// TIA Portal project "Process visualization with HMI" (V15.1) (continued)
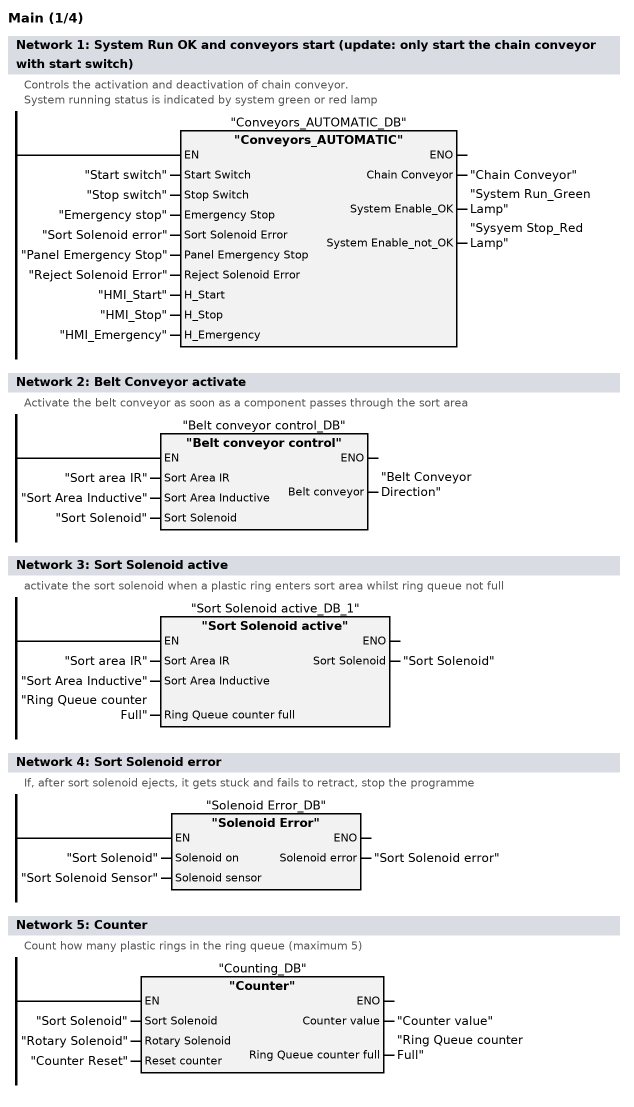
   RUNG wire#powerrail
      "Conveyors_AUTOMATIC_DB"("Start Switch" := "Start switch", "Stop Switch" := "Stop switch", "Emergency Stop" := "Emergency stop", "Sort Solenoid Error" := "Sort Solenoid error", "Panel Emergency Stop" := "Panel Emergency Stop", "Reject Solenoid Error" := "Reject Solenoid Error", H_Start := "HMI_Start", H_Stop := "HMI_Stop", H_Emergency := "HMI_Emergency", "Chain Conveyor" => "Chain Conveyor", "System Enable_OK" => "System Run_Green Lamp", "System Enable_not_OK" => "Sysyem Stop_Red Lamp")
   END_RUNG
   // the same network as SCL:
   "Conveyors_AUTOMATIC_DB"("Start Switch" := "Start switch",   // "Conveyors_AUTOMATIC"
                           "Stop Switch" := "Stop switch",
                           "Emergency Stop" := "Emergency stop",
                           "Sort Solenoid Error" := "Sort Solenoid error",
                           "Panel Emergency Stop" := "Panel Emergency Stop",
                           "Reject Solenoid Error" := "Reject Solenoid Error",
                           H_Start := "HMI_Start",
                           H_Stop := "HMI_Stop",
                           H_Emergency := "HMI_Emergency",
                           "Chain Conveyor" => "Chain Conveyor",
                           "System Enable_OK" => "System Run_Green Lamp",
                           "System Enable_not_OK" => "Sysyem Stop_Red Lamp");
END_REGION

REGION Network 2: Belt Conveyor activate
   // Activate the belt conveyor as soon as a component passes through the sort area
   RUNG wire#powerrail
      "Belt conveyor control_DB"("Sort Area IR" := "Sort area IR", "Sort Area Inductive" := "Sort Area Inductive", "Sort Solenoid" := "Sort Solenoid", "Belt conveyor" => "Belt Conveyor Direction")
   END_RUNG
   // the same network as SCL:
   "Belt conveyor control_DB"("Sort Area IR" := "Sort area IR",   // "Belt conveyor control"
                           "Sort Area Inductive" := "Sort Area Inductive",
                           "Sort Solenoid" := "Sort Solenoid",
                           "Belt conveyor" => "Belt Conveyor Direction");
END_REGION

REGION Network 3: Sort Solenoid active
   // activate the sort solenoid when a plastic ring enters sort area whilst ring queue not full
   RUNG wire#powerrail
      "Sort Solenoid active_DB_1"("Sort Area IR" := "Sort area IR", "Sort Area Inductive" := "Sort Area Inductive", "Ring Queue counter full" := "Ring Queue counter Full", "Sort Solenoid" => "Sort Solenoid")
   END_RUNG
   // the same network as SCL:
   "Sort Solenoid active_DB_1"("Sort Area IR" := "Sort area IR",   // "Sort Solenoid active"
                           "Sort Area Inductive" := "Sort Area Inductive",
                           "Ring Queue counter full" := "Ring Queue counter Full",
                           "Sort Solenoid" => "Sort Solenoid");
END_REGION

REGION Network 4: Sort Solenoid error
   // If, after sort solenoid ejects, it gets stuck and fails to retract, stop the programme
   RUNG wire#powerrail
      "Solenoid Error_DB"("Solenoid on" := "Sort Solenoid", "Solenoid sensor" := "Sort Solenoid Sensor", "Solenoid error" => "Sort Solenoid error")
   END_RUNG
   // the same network as SCL:
   "Solenoid Error_DB"("Solenoid on" := "Sort Solenoid",   // "Solenoid Error"
                       "Solenoid sensor" := "Sort Solenoid Sensor",
                       "Solenoid error" => "Sort Solenoid error");
END_REGION

REGION Network 5: Counter
   // Count how many plastic rings in the ring queue (maximum 5)
   RUNG wire#powerrail
      "Counting_DB"("Sort Solenoid" := "Sort Solenoid", "Rotary Solenoid" := "Rotary Solenoid", "Reset counter" := "Counter Reset", "Counter value" => "Counter value", "Ring Queue counter full" => "Ring Queue counter Full")
   END_RUNG
   // the same network as SCL:
   "Counting_DB"("Sort Solenoid" := "Sort Solenoid",   // "Counter"
                 "Rotary Solenoid" := "Rotary Solenoid",
                 "Reset counter" := "Counter Reset",
                 "Counter value" => "Counter value",
                 "Ring Queue counter full" => "Ring Queue counter Full");
END_REGION

REGION Network 6: Rotary Solenoid
   // activates rotary solenoid and drops plastic ring in assembly chute
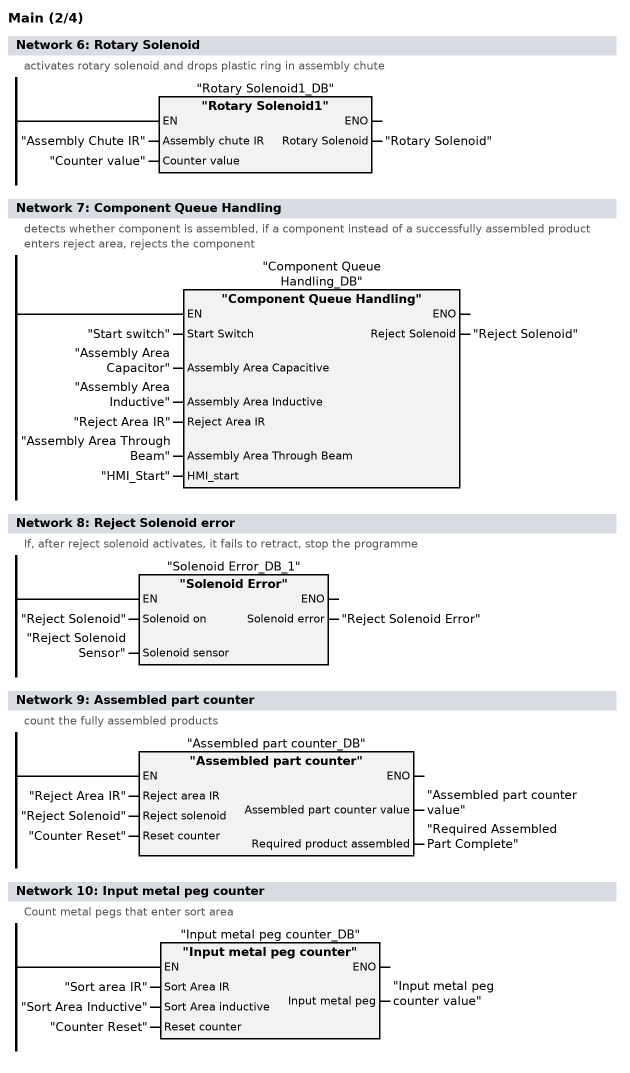
   RUNG wire#powerrail
      "Rotary Solenoid1_DB"("Assembly chute IR" := "Assembly Chute IR", "Counter value" := "Counter value", "Rotary Solenoid" => "Rotary Solenoid")
   END_RUNG
   // the same network as SCL:
   "Rotary Solenoid1_DB"("Assembly chute IR" := "Assembly Chute IR",   // "Rotary Solenoid1"
                         "Counter value" := "Counter value",
                         "Rotary Solenoid" => "Rotary Solenoid");
END_REGION

REGION Network 7: Component Queue Handling
   // detects whether component is assembled, if a component instead of a successfully assembled product enters reject area, rejects the component
   RUNG wire#powerrail
      "Component Queue Handling_DB"("Start Switch" := "Start switch", "Assembly Area Capacitive" := "Assembly Area Capacitor", "Assembly Area Inductive" := "Assembly Area Inductive", "Reject Area IR" := "Reject Area IR", "Assembly Area Through Beam" := "Assembly Area Through Beam", HMI_start := "HMI_Start", "Reject Solenoid" => "Reject Solenoid")
   END_RUNG
   // the same network as SCL:
   "Component Queue Handling_DB"("Start Switch" := "Start switch",   // "Component Queue Handling"
                           "Assembly Area Capacitive" := "Assembly Area Capacitor",
                           "Assembly Area Inductive" := "Assembly Area Inductive",
                           "Reject Area IR" := "Reject Area IR",
                           "Assembly Area Through Beam" := "Assembly Area Through Beam",
                           HMI_start := "HMI_Start",
                           "Reject Solenoid" => "Reject Solenoid");
END_REGION

REGION Network 8: Reject Solenoid error
   // If, after reject solenoid activates, it fails to retract, stop the programme
   RUNG wire#powerrail
      "Solenoid Error_DB_1"("Solenoid on" := "Reject Solenoid", "Solenoid sensor" := "Reject Solenoid Sensor", "Solenoid error" => "Reject Solenoid Error")
   END_RUNG
   // the same network as SCL:
   "Solenoid Error_DB_1"("Solenoid on" := "Reject Solenoid",   // "Solenoid Error"
                         "Solenoid sensor" := "Reject Solenoid Sensor",
                         "Solenoid error" => "Reject Solenoid Error");
END_REGION

REGION Network 9: Assembled part counter
   // count the fully assembled products
   RUNG wire#powerrail
      "Assembled part counter_DB"("Reject area IR" := "Reject Area IR", "Reject solenoid" := "Reject Solenoid", "Reset counter" := "Counter Reset", "Assembled part counter value" => "Assembled part counter value", "Required product assembled" => "Required Assembled Part Complete")
   END_RUNG
   // the same network as SCL:
   "Assembled part counter_DB"("Reject area IR" := "Reject Area IR",   // "Assembled part counter"
                           "Reject solenoid" := "Reject Solenoid",
                           "Reset counter" := "Counter Reset",
                           "Assembled part counter value" => "Assembled part counter value",
                           "Required product assembled" => "Required Assembled Part Complete");
END_REGION

REGION Network 10: Input metal peg counter
   // Count metal pegs that enter sort area
   RUNG wire#powerrail
      "Input metal peg counter_DB"("Sort Area IR" := "Sort area IR", "Sort Area inductive" := "Sort Area Inductive", "Reset counter" := "Counter Reset", "Input metal peg" => "Input metal peg counter value")
   END_RUNG
   // the same network as SCL:
   "Input metal peg counter_DB"("Sort Area IR" := "Sort area IR",   // "Input metal peg counter"
                           "Sort Area inductive" := "Sort Area Inductive",
                           "Reset counter" := "Counter Reset",
                           "Input metal peg" => "Input metal peg counter value");
END_REGION

REGION Network 11: Input plastic ring counter
   // Count plastic ring that enters sort area
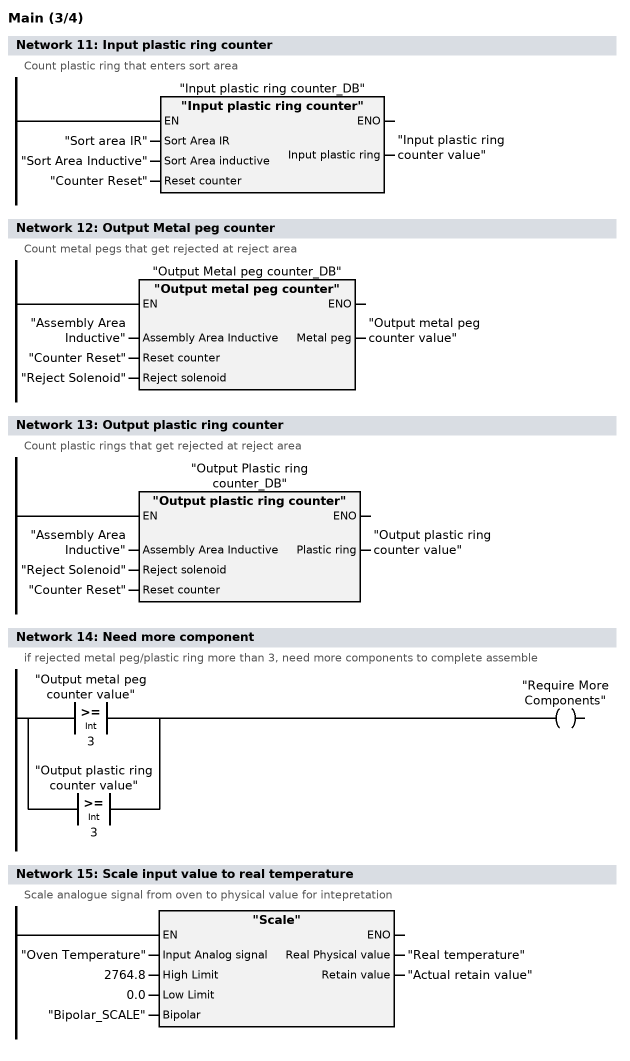
   RUNG wire#powerrail
      "Input plastic ring counter_DB"("Sort Area IR" := "Sort area IR", "Sort Area inductive" := "Sort Area Inductive", "Reset counter" := "Counter Reset", "Input plastic ring" => "Input plastic ring counter value")
   END_RUNG
   // the same network as SCL:
   "Input plastic ring counter_DB"("Sort Area IR" := "Sort area IR",   // "Input plastic ring counter"
                           "Sort Area inductive" := "Sort Area Inductive",
                           "Reset counter" := "Counter Reset",
                           "Input plastic ring" => "Input plastic ring counter value");
END_REGION

REGION Network 12: Output Metal peg counter
   // Count metal pegs that get rejected at reject area
   RUNG wire#powerrail
      "Output Metal peg counter_DB"("Assembly Area Inductive" := "Assembly Area Inductive", "Reset counter" := "Counter Reset", "Reject solenoid" := "Reject Solenoid", "Metal peg" => "Output metal peg counter value")
   END_RUNG
   // the same network as SCL:
   "Output Metal peg counter_DB"("Assembly Area Inductive" := "Assembly Area Inductive",   // "Output metal peg counter"
                           "Reset counter" := "Counter Reset",
                           "Reject solenoid" := "Reject Solenoid",
                           "Metal peg" => "Output metal peg counter value");
END_REGION

REGION Network 13: Output plastic ring counter
   // Count plastic rings that get rejected at reject area
   RUNG wire#powerrail
      "Output Plastic ring counter_DB"("Assembly Area Inductive" := "Assembly Area Inductive", "Reject solenoid" := "Reject Solenoid", "Reset counter" := "Counter Reset", "Plastic ring" => "Output plastic ring counter value")
   END_RUNG
   // the same network as SCL:
   "Output Plastic ring counter_DB"("Assembly Area Inductive" := "Assembly Area Inductive",   // "Output plastic ring counter"
                           "Reject solenoid" := "Reject Solenoid",
                           "Reset counter" := "Counter Reset",
                           "Plastic ring" => "Output plastic ring counter value");
END_REGION

REGION Network 14: Need more component
   // if rejected metal peg/plastic ring more than 3, need more components to complete assemble
   RUNG wire#powerrail
      { S7_Templates := "SrcType := Int" } GE_Contact(in1 := "Output metal peg counter value", in2 := 3)
      wire#w1
      Coil( "Require More Components" )
   END_RUNG
   RUNG wire#powerrail
      { S7_Templates := "SrcType := Int" } GE_Contact(in1 := "Output plastic ring counter value", in2 := 3)
   END_RUNG wire#w1
   // the same network as SCL:
   "Require More Components" := ("Output metal peg counter value" >= 3) OR ("Output plastic ring counter value" >= 3);
END_REGION

REGION Network 15: Scale input value to real temperature
   // Scale analogue signal from oven to physical value for intepretation
   RUNG wire#powerrail
      "Scale"("Input Analog signal" := "Oven Temperature", "High Limit" := 2764.8, "Low Limit" := 0.0, Bipolar := "Bipolar_SCALE", "Real Physical value" => "Real temperature", "Retain value" => "Actual retain value")
   END_RUNG
   // the same network as SCL:
   "Scale"("Input Analog signal" := "Oven Temperature",
           "High Limit" := 2764.8,
           "Low Limit" := 0.0,
           Bipolar := "Bipolar_SCALE",
           "Real Physical value" => "Real temperature",
           "Retain value" => "Actual retain value");
END_REGION

REGION Network 16: Unscale
   // scale physical temperature value back to analogue signal
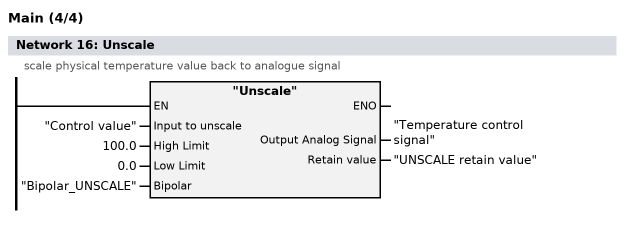
   RUNG wire#powerrail
      "Unscale"("Input to unscale" := "Control value", "High Limit" := 100.0, "Low Limit" := 0.0, Bipolar := "Bipolar_UNSCALE", "Output Analog Signal" => "Temperature control signal", "Retain value" => "UNSCALE retain value")
   END_RUNG
   // the same network as SCL:
   "Unscale"("Input to unscale" := "Control value",
             "High Limit" := 100.0,
             "Low Limit" := 0.0,
             Bipolar := "Bipolar_UNSCALE",
             "Output Analog Signal" => "Temperature control signal",
             "Retain value" => "UNSCALE retain value");
END_REGION
END_ORGANIZATION_BLOCK

ORGANIZATION_BLOCK "Cyclic interrupt"   // OB30, LAD, CyclicInterrupt
TITLE = PID Controller
{ S7_Optimized_Access := 'TRUE' }
VERSION : 0.1
   VAR_INPUT
      Initial_Call : Bool;   // Initial call of this OB
      Event_Count : Int;   // Events discarded
   END_VAR
BEGIN

REGION Network 1: PID control for oven temperature
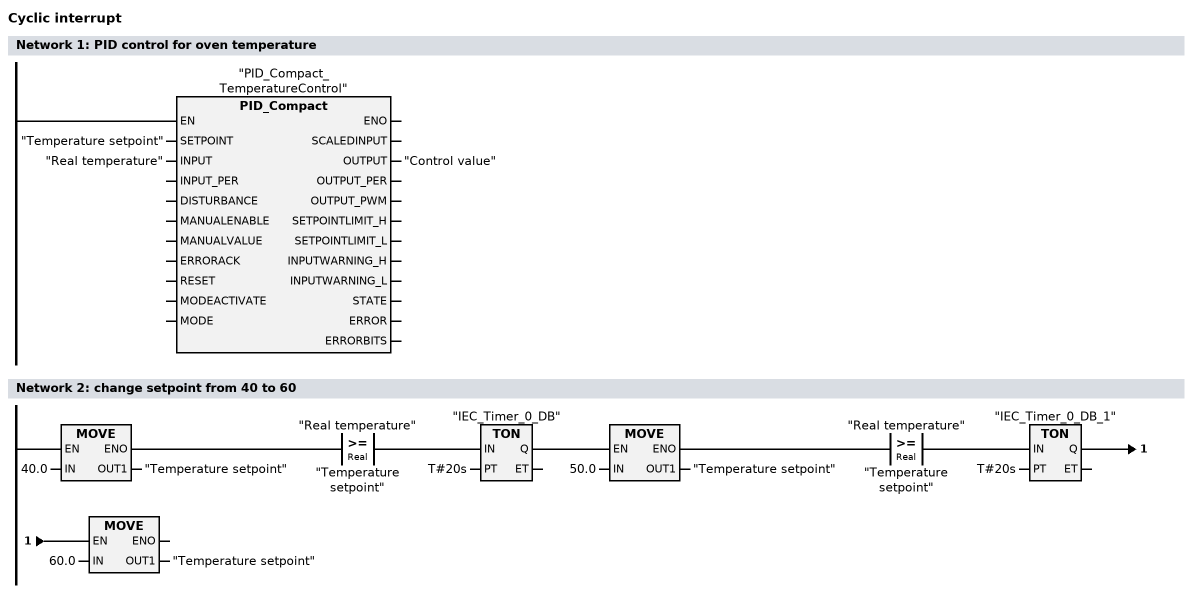
   "PID_Compact_TemperatureControl"(Setpoint := "Temperature setpoint",   // PID_Compact
                           Input := "Real temperature",
                           Output => "Control value");
END_REGION

REGION Network 2: change setpoint from 40 to 60
   "Temperature setpoint" := 40.0;
   "IEC_Timer_0_DB".TON(IN := "Real temperature" >= "Temperature setpoint", PT := T#20s);
   IF "IEC_Timer_0_DB".Q THEN "Temperature setpoint" := 50.0; END_IF;
   "IEC_Timer_0_DB_1".TON(IN := "IEC_Timer_0_DB".Q AND ("Real temperature" >= "Temperature setpoint"),
                          PT := T#20s);
   IF "IEC_Timer_0_DB_1".Q THEN "Temperature setpoint" := 60.0; END_IF;
END_REGION

REGION Network 3: change setpoint from 60 to 50
END_REGION
END_ORGANIZATION_BLOCK

(* ===== HMI "HMI_RT_1" =====
system functions are stored by id; their names below are inferred from use
connection "HMI_Connection_1": ETHERNET, S7_1500_OMS

HMI tags "Default tag table"
   "Counter value" : Int = PLC "Counter value" AT %MW0, 100 ms
   "Sort Solenoid Sensor" : Bool = PLC "Sort Solenoid Sensor" AT %I0.6, 100 ms
   "Counter Reset" : Bool = PLC "Counter Reset" AT %M4.4, 100 ms
   "HMI_Stop" : Bool = PLC HMI_Stop AT %M4.2, 100 ms
   "HMI_Start" : Bool = PLC HMI_Start AT %M4.1, 100 ms
   "Emergency stop" : Bool = PLC "Emergency stop" AT %I1.0, 100 ms
   "Stop switch" : Bool = PLC "Stop switch" AT %I0.3, 100 ms
   "System Run_Green Lamp" : Bool = PLC "System Run_Green Lamp" AT %Q3.0, 100 ms
   "Sysyem Stop_Red Lamp" : Bool = PLC "Sysyem Stop_Red Lamp" AT %Q3.2, 100 ms
   "Chain Conveyor" : Bool = PLC "Chain Conveyor" AT %Q0.0, 100 ms
   "Sort area IR" : Bool = PLC "Sort area IR" AT %I0.4, 100 ms
   "Sort Area Inductive" : Bool = PLC "Sort Area Inductive" AT %I0.5, 100 ms
   "Assembly Area Inductive" : Bool = PLC "Assembly Area Inductive" AT %I1.3, 100 ms
   "Assembly Area Capacitor" : Bool = PLC "Assembly Area Capacitor" AT %I1.2, 100 ms
   "Assembly Chute IR" : Bool = PLC "Assembly Chute IR" AT %I0.7, 100 ms
   "Reject Solenoid" : Bool = PLC "Reject Solenoid" AT %Q0.2, 100 ms
   "Reject Solenoid Sensor" : Bool = PLC "Reject Solenoid Sensor" AT %I1.5, 100 ms
   "Belt Conveyor Direction" : Bool = PLC "Belt Conveyor Direction" AT %Q0.4, 100 ms
   "Assembly Area Through Beam" : Bool = PLC "Assembly Area Through Beam" AT %I1.1, 100 ms
   "Assembled part counter value" : Int = PLC "Assembled part counter value" AT %MW40, 100 ms
   "Input metal peg counter value" : Int = PLC "Input metal peg counter value" AT %MW80, 100 ms
   "Input plastic ring counter value" : Int = PLC "Input plastic ring counter value" AT %MW100, 100 ms
   "Output metal peg counter value" : Int = PLC "Output metal peg counter value" AT %MW50, 100 ms
   "Output plastic ring counter value" : Int = PLC "Output plastic ring counter value" AT %MW60, 100 ms
   "Ring Queue counter Full" : Bool = PLC "Ring Queue counter Full" AT %M4.0, 100 ms
   "HMI_Emergency" : Bool = PLC HMI_Emergency AT %M4.5, 100 ms
   "Panel Emergency Stop" : Bool = PLC "Panel Emergency Stop" AT %I2.7, 100 ms
   "Real temperature" : Real = PLC "Real temperature" AT %MD5, 100 ms
   "ON/OFF Temperature set point" : Real = PLC "ON/OFF Temperature set point" AT %MD20, 100 ms
   "Required Assembled Part Complete" : Bool = PLC "Required Assembled Part Complete" AT %M9.0, 100 ms
   "Require More Components" : Bool = PLC "Require More Components" AT %M9.1, 100 ms

Template "Template_1" 800x480
   Button "Exit" at 720,420 size 78x58; TextOff 'Exit'; PictureOff "ExitRuntime_TP700_Comfort_TR"; PictureOn "ExitRuntime_TP700_Comfort_TR"
      on Release: StopRuntime(0)
   Button "Template_Button" at 640,420 size 78x58; TextOff 'Text'
   Button "Template_Button_1" at 560,420 size 78x58; TextOff 'Text'
   Button "Template_Button_2" at 480,420 size 78x58; TextOff 'Text'
   Button "Template_Button_3" at 400,420 size 78x58; TextOff 'Text'
   Button "Template_Button_4" at 321,420 size 78x58; TextOff 'Text'
   Button "Template_Button_5" at 241,420 size 78x58; TextOff 'Text'
   Button "Template_Button_6" at 161,420 size 78x58; TextOff 'Text'
   Button "Template_Button_7" at 81,420 size 78x58; TextOff 'Text'
   Button "Start screen" at 1,420 size 78x58; TextOff 'Start screen'; PictureOff "NavigateHome_TP700_Comfort_TR"; PictureOn "NavigateHome_TP700_Comfort_TR"
      on Release: ActivateScreen("Sorting Station Overview", 0)

screen "Sorting Station Overview" 800x480, template "Template_1"
   TextField "HmiScreenItemData_5" at 80,196 size 640x25; Text 'Welcome to HMI_1 (TP700 Comfort)!'
   Button "HmiScreenItemData" at 36,36 size 159x47; TextOff 'System Control'; PictureOff "Navigates to System Control for TP700 Comfort 15.1.0.0"; PictureOn "Navigates to System Control for TP700 Comfort 15.1.0.0"
      on Release: ActivateScreen("System Control", 0)
   Button "HmiScreenItemData_1" at 36,95 size 159x47; TextOff 'Input/Output'; PictureOff "Navigates to Input/Output for TP700 Comfort 15.1.0.0"; PictureOn "Navigates to Input/Output for TP700 Comfort 15.1.0.0"
      on Release: ActivateScreen("Input/Output", 0)
   Button "HmiScreenItemData_2" at 36,154 size 159x47; TextOff 'Temperature Control'; PictureOff "Navigates to Temperature Control for TP700 Comfort 15.1.0.0"; PictureOn "Navigates to Temperature Control for TP700 Comfort 15.1.0.0"
      on Release: ActivateScreen("Temperature Control", 0)
   Button "HmiScreenItemData_3" at 36,213 size 159x47; TextOff 'Alarm'; PictureOff "Navigates to Alarm for TP700 Comfort 15.1.0.0"; PictureOn "Navigates to Alarm for TP700 Comfort 15.1.0.0"
      on Release: ActivateScreen("Alarm", 0)
   Button "HmiScreenItemData_4" at 36,272 size 159x47; TextOff 'Exercise'; PictureOff "Navigates to Exercise for TP700 Comfort 15.1.0.0"; PictureOn "Navigates to Exercise for TP700 Comfort 15.1.0.0"
      on Release: ActivateScreen("Exercise", 0)
   Button "HmiScreenItemData_6" at 36,331 size 159x47; TextOff 'System screens'; PictureOff "Navigates to System screens for TP700 Comfort 15.1.0.0"; PictureOn "Navigates to System screens for TP700 Comfort 15.1.0.0"
      on Release: ActivateScreen("System screens", 0)
   GraphicView "Graphic view_1" at 230,64 size 473x289; Picture "HMI picture"
   Button "HmiScreenItemData_7" at 212,15 size 159x47; TextOn 'ON/OFF Control'; TextOff 'ON/OFF Control'; PictureOn "Navigates to System screens for TP700 Comfort 15.1.0.0"; PictureOff "Navigates to System screens for TP700 Comfort 15.1.0.0"
      on Release: ActivateScreen("ON/OFF Control", 0)

screen "System Control" 800x480, template "Template_1"
   Button "Back" at 1,1 size 159x47; TextOff 'Back'
      on Release: ActivateScreen("Sorting Station Overview", 0)
   GraphicView "Graphic view_1" at 0,0 size 800x480; Picture "bytronic"
   Button "Back_1" at 0,28 size 159x47; TextOn 'Back'; TextOff 'Back'
      on Release: ActivateScreen("Sorting Station Overview", 0)
   IOField "I/O field_1" at 23,335 size 29x32; FormatPattern 9
      ProcessValue <- "Counter value"
   TextField "Text field_1" at 6,303 size 124x23; Text 'Counter Value'
   Circle "Circle_1" at 241,32 size 18x18
      Appearance <- "Sort Solenoid Sensor"
   Circle "Circle_2" at 65,331 size 35x35
      Appearance <- "Ring Queue counter Full"
   Button "Button_1" at 283,412 size 40x40; TextOff 'Text'; PictureOn "Pushbutton_Round_R_On_256c"; PictureOff "Pushbutton_Round_R_Off_256c"
      on Press: function_b14e0dd5("Counter Reset", 0)
   Button "Button_2" at 139,412 size 40x40; TextOff 'Text'; PictureOn "Pushbutton_Round_R_On_256c"; PictureOff "Pushbutton_Round_R_Off_256c"
      on Press: function_b14e0dd5("HMI_Stop", 0)
   Button "Button_3" at 182,412 size 40x40; TextOff 'Text'; PictureOn "Pushbutton_Round_G_On_256c"; PictureOff "Pushbutton_Round_G_Off_256c"
      on Press: function_b14e0dd5("HMI_Start", 0)
   Circle "Circle_3" at 240,108 size 20x20
      Appearance <- "Sort Area Inductive"
   Circle "Circle_4" at 418,387 size 25x25
      Appearance <- "Sysyem Stop_Red Lamp"
   Circle "Circle_5" at 418,413 size 25x25
      Appearance <- "HMI_Emergency"
   Circle "Circle_6" at 418,439 size 25x25
      Appearance <- "System Run_Green Lamp"
   Rectangle "Rectangle_1" at 131,153 size 28x18
      Appearance <- "Chain Conveyor"
   Rectangle "Rectangle_2" at 224,101 size 9x24
      Appearance <- "Sort area IR"
   Rectangle "Rectangle_3" at 308,218 size 27x19
      Appearance <- "Assembly Area Capacitor"
   Circle "Circle_7" at 313,275 size 18x18
      Appearance <- "Assembly Area Inductive"
   Rectangle "Rectangle_4" at 241,295 size 18x10
      Appearance <- "Assembly Chute IR"
   Circle "Circle_8" at 498,347 size 16x16
      Appearance <- "Reject Solenoid Sensor"
   Rectangle "Rectangle_5" at 519,334 size 19x25
      Appearance <- "Belt Conveyor Direction"
   Circle "Circle_9" at 343,253 size 14x14
      Appearance <- "Assembly Area Through Beam"
   IOField "I/O field_2" at 728,378 size 63x25; FormatPattern 999
      ProcessValue <- "Assembled part counter value"
   Switch "Switch_1" at 6,377 size 100x100; CaptionText 'Switch'; TextOff 'OFF'; TextOn 'ON'; PictureOn "Pushbutton_Emergency_On_256c"; PictureOff "Pushbutton_Emergency_Off_256c"
      ProcessValue <- "HMI_Emergency"
   IOField "I/O field_3" at 653,378 size 63x25; FormatPattern 999
      ProcessValue <- "Output metal peg counter value"
   IOField "I/O field_4" at 576,378 size 63x25; FormatPattern 999
      ProcessValue <- "Output plastic ring counter value"
   TextField "Text field_2" at 285,33 size 504x23; Text 'All the required products have been assembled !'
      Appearance <- "Required Assembled Part Complete"
   TextField "Text field_4" at 285,48 size 350x42; Text 'Process cannot be completed, and more products should be ordered.'
      Appearance <- "Require More Components"

screen "Input/Output" 800x480, template "Template_1"
   Button "Back" at 1,1 size 159x47; TextOff 'Back'
      on Release: ActivateScreen("Sorting Station Overview", 0)
   TextField "Text field_1" at 43,63 size 143x23; Text 'Counter Value'
   TextField "Text field_2" at 249,48 size 70x23; Text 'Inputs'
   TextField "Text field_3" at 544,48 size 76x23; Text 'Outputs'
   Bar "Bar_1" at 63,104 size 80x230; MinimumValue 0
      ProcessValue <- "Counter value"
   Bar "Bar_2" at 650,113 size 80x230; MinimumValue 0; MaximumValue 100
      ProcessValue <- "Assembled part counter value"
   TextField "Text field_4" at 619,78 size 165x23; Text 'Assembled Parts'
   IOField "I/O field_1" at 440,289 size 69x32; FormatPattern 999
      ProcessValue <- "Assembled part counter value"
   TextField "Text field_5" at 431,89 size 100x23; Text 'Metal peg'
   TextField "Text field_6" at 422,174 size 115x23; Text 'Plastic ring'
   IOField "I/O field_2" at 440,208 size 69x32; FormatPattern 999
      ProcessValue <- "Output plastic ring counter value"
   IOField "I/O field_3" at 440,123 size 69x32; FormatPattern 999
      ProcessValue <- "Output metal peg counter value"
   TextField "Text field_7" at 407,260 size 164x23; Text 'Assembled Parts'
   TextField "Text field_8" at 233,108 size 100x23; Text 'Metal peg'
   TextField "Text field_9" at 233,244 size 115x23; Text 'Plastic ring'
   IOField "I/O field_4" at 245,274 size 69x32; FormatPattern 999
      ProcessValue <- "Input plastic ring counter value"
   IOField "I/O field_5" at 245,153 size 69x32; FormatPattern 999
      ProcessValue <- "Input metal peg counter value"
   Rectangle "Rectangle_1" at 75,392 size 50x30
      Appearance <- "Chain Conveyor"
   TextField "Text field_10" at 38,354 size 143x23; Text 'Chain conveyor'
   TextField "Text field_11" at 219,355 size 129x23; Text 'Belt conveyor'
   Rectangle "Rectangle_2" at 253,392 size 50x30
      Appearance <- "Belt Conveyor Direction"
   TextField "Text field_12" at 294,14 size 506x23; Text 'For sensors info, please refer to "System Control" page'
   Circle "Circle_1" at 415,407 size 34x34
      Appearance <- "Emergency stop"
   Circle "Circle_2" at 671,390 size 34x34
      Appearance <- "Panel Emergency Stop"
   TextField "Text field_13" at 407,345 size 150x23; Text 'Emergency Stop'
   TextField "Text field_14" at 619,354 size 160x23; Text 'Panel Emergency'
   Circle "Circle_3" at 509,407 size 34x34
      Appearance <- "HMI_Emergency"
   TextField "Text field_15" at 401,377 size 85x23; Text 'Physical'
   TextField "Text field_16" at 505,377 size 41x23; Text 'HMI'

screen "Temperature Control" 800x480, template "Template_1"
   TextField "HmiScreenItemData" at 80,196 size 640x25; Text 'Temperature Control'
   Button "Back" at 1,1 size 159x47; TextOff 'Back'
      on Release: ActivateScreen("Sorting Station Overview", 0)

screen "Alarm" 800x480, template "Template_1"
   TextField "HmiScreenItemData" at 80,196 size 640x25; Text 'Alarm'
   Button "Back" at 1,1 size 159x47; TextOff 'Back'
      on Release: ActivateScreen("Sorting Station Overview", 0)

screen "Exercise" 800x480, template "Template_1"
   TextField "HmiScreenItemData" at 80,196 size 640x25; Text 'Exercise'
   Button "Back" at 1,1 size 159x47; TextOff 'Back'
      on Release: ActivateScreen("Sorting Station Overview", 0)

screen "System screens" 800x480, template "Template_1"
   Button "Back" at 1,1 size 159x47; TextOff 'Back'
      on Release: ActivateScreen("Sorting Station Overview", 0)
   Button "HmiScreenItemData" at 36,95 size 159x47; TextOff 'SIMATIC PLC system diagnos...'; PictureOff "Navigates to SIMATIC PLC system diagnostics for TP700 Comfort 15.1.0.0"; PictureOn "Navigates to SIMATIC PLC system diagnostics for TP700 Comfort 15.1.0.0"
      on Release: ActivateScreen("SIMATIC PLC system diagnostics", 0)

screen "SIMATIC PLC system diagnostics" 800x480, template "Template_1"
   SysDiagControl "HmiScreenItemData" at 1,49 size 796x364
   Button "Back" at 1,1 size 159x47; TextOff 'Back'
      on Release: ActivateScreen("System screens", 0)

screen "ON/OFF Control" 800x480
   Button "Back" at 1,1 size 159x47; TextOn 'Back'; TextOff 'Back'
      on Release: ActivateScreen("Sorting Station Overview", 0)
   TrendView "Trend view_1" at 158,1 size 642x479
   IOField "I/O field_1" at 37,360 size 64x32; FormatPattern 999.9
      ProcessValue <- "ON/OFF Temperature set point"
   Bar "Bar_1" at 27,113 size 80x230; MinimumValue 0; MaximumValue 100
      ProcessValue <- "ON/OFF Temperature set point"
   TextField "Text field_1" at 30,60 size 72x23; Text 'On/Off'
   TextField "Text field_2" at 1,83 size 144x23; Text 'Temp Set point'
*)